REGION Network 6
   RUNG wire#powerrail
      "FB_CONCAT_STRINGS_FOR_MQTT_DB"(temperature1 := "DB_GlobalData".RTDs.RTD1.ch0, temperature2 := "DB_GlobalData".RTDs.RTD1.ch1, temperature3 := "DB_GlobalData".RTDs.RTD1.ch2, temperature4 := "DB_GlobalData".RTDs.RTD1.ch3, strCombinedString => "MQTT_DB".MQTT_CLIEENTS[0].mqttUserControl.sStringToPublish, q_aStringToSendToMqtt =>)
      "FB_CONCAT_STRINGS_FOR_MQTT_1_DB"(temperature1 := "DB_GlobalData".RTDs.RTD1.ch0, temperature2 := "DB_GlobalData".RTDs.RTD1.ch1, temperature3 :=, temperature4 := "DB_GlobalData".RTDs.RTD1.ch2, customText := '', strCombinedString =>, q_aStringToSendToMqtt => "MQTT_DB".MQTT_CLIENTS_WSTRING[0].mqttParam.message)
   END_RUNG
   // the same network as SCL:
   "FB_CONCAT_STRINGS_FOR_MQTT_DB"(temperature1 := "DB_GlobalData".RTDs.RTD1.ch0,   // "FB_CONCAT_STRINGS_FOR_MQTT"
                           temperature2 := "DB_GlobalData".RTDs.RTD1.ch1,
                           temperature3 := "DB_GlobalData".RTDs.RTD1.ch2,
                           temperature4 := "DB_GlobalData".RTDs.RTD1.ch3,
                           strCombinedString => "MQTT_DB".MQTT_CLIEENTS[0].mqttUserControl.sStringToPublish,
                           ENO => #_w1);
   IF #_w1 THEN
       "FB_CONCAT_STRINGS_FOR_MQTT_1_DB"(temperature1 := "DB_GlobalData".RTDs.RTD1.ch0,   // "FB_CONCAT_STRINGS_FOR_MQTT_1"
                               temperature2 := "DB_GlobalData".RTDs.RTD1.ch1,
                               temperature4 := "DB_GlobalData".RTDs.RTD1.ch2,
                               customText := '',
                               q_aStringToSendToMqtt => "MQTT_DB".MQTT_CLIENTS_WSTRING[0].mqttParam.message);
   END_IF;
END_REGION

REGION Network 7: MQTT publisher 1
   RUNG wire#powerrail
      "LMqtt_Publisher_DB1"(publish := wire#w1, enable := "MQTT_DB".MQTT_CLIEENTS[0].mqttUserControl.xEnable, tcpConnParam := "MQTT_DB".MQTT_CLIEENTS[0].mqttTcpParam, mqttParam := "MQTT_DB".MQTT_CLIEENTS[0].mqttParam, tcpEstablished => "MQTT_DB".MQTT_CLIEENTS[0].mqttUserControl.Status.xtcpEsablished, mqttEstablished => "MQTT_DB".MQTT_CLIEENTS[0].mqttUserControl.Status.xmqttEstavlished, published => "MQTT_DB".MQTT_CLIEENTS[0].mqttUserControl.Status.xpublished, busy => "MQTT_DB".MQTT_CLIEENTS[0].mqttUserControl.Status.xbusy, error => "MQTT_DB".MQTT_CLIEENTS[0].mqttUserControl.Status.xerror, status => "MQTT_DB".MQTT_CLIEENTS[0].mqttUserControl.Status.status, statusID => "MQTT_DB".MQTT_CLIEENTS[0].mqttUserControl.Status.istatusID)
   END_RUNG
   RUNG wire#powerrail
      Contact( "MQTT_DB".MQTT_CLIEENTS[0].mqttUserControl.xPusblish )
   END_RUNG wire#w1
   // the same network as SCL:
   "LMqtt_Publisher_DB1"(enable := "MQTT_DB".MQTT_CLIEENTS[0].mqttUserControl.xEnable,   // "LMqtt_Publisher"
                         publish := "MQTT_DB".MQTT_CLIEENTS[0].mqttUserControl.xPusblish,
                         tcpConnParam := "MQTT_DB".MQTT_CLIEENTS[0].mqttTcpParam,
                         mqttParam := "MQTT_DB".MQTT_CLIEENTS[0].mqttParam,
                         tcpEstablished => "MQTT_DB".MQTT_CLIEENTS[0].mqttUserControl.Status.xtcpEsablished,
                         mqttEstablished => "MQTT_DB".MQTT_CLIEENTS[0].mqttUserControl.Status.xmqttEstavlished,
                         published => "MQTT_DB".MQTT_CLIEENTS[0].mqttUserControl.Status.xpublished,
                         busy => "MQTT_DB".MQTT_CLIEENTS[0].mqttUserControl.Status.xbusy,
                         error => "MQTT_DB".MQTT_CLIEENTS[0].mqttUserControl.Status.xerror,
                         status => "MQTT_DB".MQTT_CLIEENTS[0].mqttUserControl.Status.status,
                         statusID => "MQTT_DB".MQTT_CLIEENTS[0].mqttUserControl.Status.istatusID);
END_REGION

REGION Network 8: MQTT-WSTRING-TEST
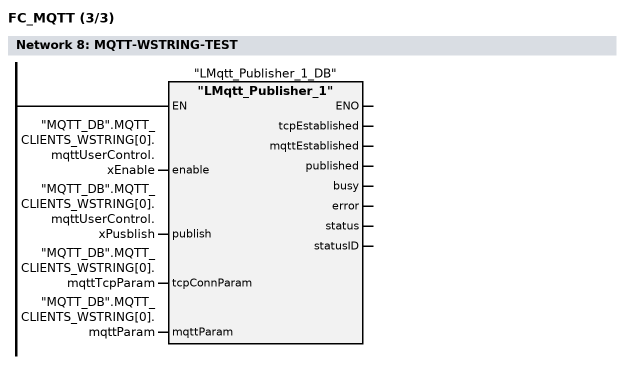
   RUNG wire#powerrail
      "LMqtt_Publisher_1_DB"(enable := "MQTT_DB".MQTT_CLIENTS_WSTRING[0].mqttUserControl.xEnable, publish := "MQTT_DB".MQTT_CLIENTS_WSTRING[0].mqttUserControl.xPusblish, tcpConnParam := "MQTT_DB".MQTT_CLIENTS_WSTRING[0].mqttTcpParam, mqttParam := "MQTT_DB".MQTT_CLIENTS_WSTRING[0].mqttParam, tcpEstablished =>, mqttEstablished =>, published =>, busy =>, error =>, status =>, statusID =>)
   END_RUNG
   // the same network as SCL:
   "LMqtt_Publisher_1_DB"(enable := "MQTT_DB".MQTT_CLIENTS_WSTRING[0].mqttUserControl.xEnable,   // "LMqtt_Publisher_1"
                          publish := "MQTT_DB".MQTT_CLIENTS_WSTRING[0].mqttUserControl.xPusblish,
                          tcpConnParam := "MQTT_DB".MQTT_CLIENTS_WSTRING[0].mqttTcpParam,
                          mqttParam := "MQTT_DB".MQTT_CLIENTS_WSTRING[0].mqttParam);
END_REGION
END_FUNCTION

FUNCTION "FC_CalculatePressRPM" : Void   // FC9, LAD
{ S7_Optimized_Access := 'TRUE' }
VERSION : 0.1
   VAR_INPUT
      i_xPulse : Bool;   // Pulse for every turn
   END_VAR
   VAR_IN_OUT
      i_iCurrentCounter : Int;
      q_iRealSPeed : Int;
   END_VAR
   VAR_TEMP
      xcalculateRPM : Bool;
      _xton : Bool;
      Temp_RPM : Real;
   END_VAR
   VAR_TEMP   // added for the SCL form of the ladder/FBD networks
      _w1 : Bool;
   END_VAR
BEGIN

REGION Network 2: 5S TIMER
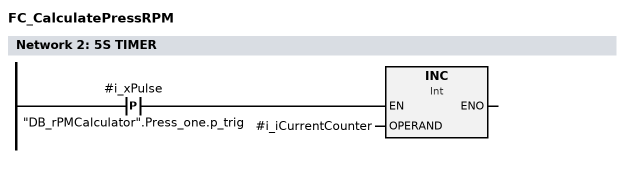
   RUNG wire#powerrail
      P_Contact(operand := #i_xPulse, bit := "DB_rPMCalculator".Press_one.p_trig)
      { S7_Templates := "DestType := Int" } Inc( #i_iCurrentCounter )
   END_RUNG
   // the same network as SCL:
   #_w1 := #i_xPulse AND NOT "DB_rPMCalculator".Press_one.p_trig;   // rising edge of #i_xPulse
   "DB_rPMCalculator".Press_one.p_trig := #i_xPulse;
   IF #_w1 THEN #i_iCurrentCounter := #i_iCurrentCounter + 1; END_IF;
END_REGION

REGION Network 3 (SCL)
   // Start 5-second timer
   "DB_rPMCalculator".Press_one.PulseTimer(IN := TRUE, PT := T#5s);



   // When 5 seconds have passed, calculate RPM
   IF "DB_rPMCalculator".Press_one.PulseTimer.Q THEN
       #q_iRealSPeed := INT_TO_REAL(#i_iCurrentCounter * 60.0) / (5.0);  // Calculate RPM
      // #q_iRealSPeed := #Temp_RPM;                      // Set the output RPM

       // Reset pulse count and timer
       #i_iCurrentCounter := 0;
       "DB_rPMCalculator".Press_one.PulseTimer(IN := FALSE,
                                               PT := T#5s);                // Reset the timer
   END_IF;
END_REGION
END_FUNCTION

FUNCTION "FC_AKD_PNU" : Void   // FC10, LAD
{ S7_Optimized_Access := 'TRUE' }
VERSION : 0.1
   VAR_INPUT
      HW_IO_telegram : Hw_Io;
   END_VAR
   VAR_IN_OUT
      AKD_PNU_v02_Instance : "AKD_PNU_v02";
      IO_DATA : "PNU_DATA";
   END_VAR
BEGIN

REGION Network 1: AKD1
   // AKD FB
   // 
   // set ID - to telegram ID of a AKD
   // 
   // 
   // # Read data from AKD PNU #
   // =================================================
   // 
   // 1. set PNU number and PNU subindex (iPNUnumber, iPNUsubindex)
   // 2. set cmd.xstartRead bit to One
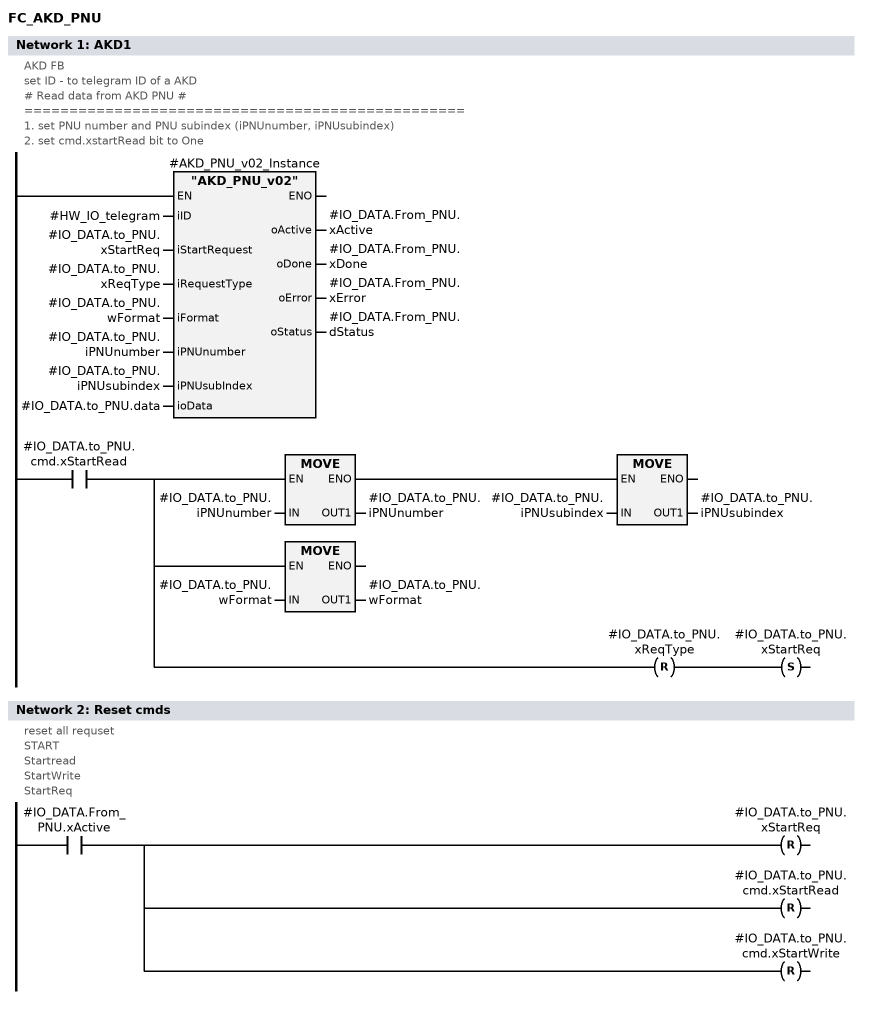
   RUNG wire#powerrail
      #AKD_PNU_v02_Instance(iID := #HW_IO_telegram, iStartRequest := #IO_DATA.to_PNU.xStartReq, iRequestType := #IO_DATA.to_PNU.xReqType, iFormat := #IO_DATA.to_PNU.wFormat, iPNUnumber := #IO_DATA.to_PNU.iPNUnumber, iPNUsubIndex := #IO_DATA.to_PNU.iPNUsubindex, ioData := #IO_DATA.to_PNU.data, oActive => #IO_DATA.From_PNU.xActive, oDone => #IO_DATA.From_PNU.xDone, oError => #IO_DATA.From_PNU.xError, oStatus => #IO_DATA.From_PNU.dStatus)
   END_RUNG
   RUNG wire#powerrail
      Contact( #IO_DATA.to_PNU.cmd.xStartRead )
      wire#w1
      Move(in := #IO_DATA.to_PNU.iPNUnumber, out1 => #IO_DATA.to_PNU.iPNUnumber)
      Move(in := #IO_DATA.to_PNU.iPNUsubindex, out1 => #IO_DATA.to_PNU.iPNUsubindex)
   END_RUNG
   RUNG wire#w1
      Move(in := #IO_DATA.to_PNU.wFormat, out1 => #IO_DATA.to_PNU.wFormat)
   END_RUNG
   RUNG wire#w1
      R_Coil( #IO_DATA.to_PNU.xReqType )
      S_Coil( #IO_DATA.to_PNU.xStartReq )
   END_RUNG
   // the same network as SCL:
   #AKD_PNU_v02_Instance(iID := #HW_IO_telegram,   // "AKD_PNU_v02"
                         iStartRequest := #IO_DATA.to_PNU.xStartReq,
                         iRequestType := #IO_DATA.to_PNU.xReqType,
                         iFormat := #IO_DATA.to_PNU.wFormat,
                         iPNUnumber := #IO_DATA.to_PNU.iPNUnumber,
                         iPNUsubIndex := #IO_DATA.to_PNU.iPNUsubindex,
                         ioData := #IO_DATA.to_PNU.data,
                         oActive => #IO_DATA.From_PNU.xActive,
                         oDone => #IO_DATA.From_PNU.xDone,
                         oError => #IO_DATA.From_PNU.xError,
                         oStatus => #IO_DATA.From_PNU.dStatus);
   IF #IO_DATA.to_PNU.cmd.xStartRead THEN
       #IO_DATA.to_PNU.iPNUnumber := #IO_DATA.to_PNU.iPNUnumber;
       #IO_DATA.to_PNU.iPNUsubindex := #IO_DATA.to_PNU.iPNUsubindex;
       #IO_DATA.to_PNU.wFormat := #IO_DATA.to_PNU.wFormat;
       #IO_DATA.to_PNU.xReqType := FALSE;
       #IO_DATA.to_PNU.xStartReq := TRUE;
   END_IF;
END_REGION

REGION Network 2: Reset cmds
   // reset all requset
   // 
   // START
   // Startread
   // StartWrite
   // StartReq
   RUNG wire#powerrail
      Contact( #IO_DATA.From_PNU.xActive )
      wire#w1
      R_Coil( #IO_DATA.to_PNU.xStartReq )
   END_RUNG
   RUNG wire#w1
      R_Coil( #IO_DATA.to_PNU.cmd.xStartRead )
   END_RUNG
   RUNG wire#w1
      R_Coil( #IO_DATA.to_PNU.cmd.xStartWrite )
   END_RUNG
   // the same network as SCL:
   IF #IO_DATA.From_PNU.xActive THEN
       #IO_DATA.to_PNU.xStartReq := FALSE;
       #IO_DATA.to_PNU.cmd.xStartRead := FALSE;
       #IO_DATA.to_PNU.cmd.xStartWrite := FALSE;
   END_IF;
END_REGION
END_FUNCTION

FUNCTION "FC_MotorControl" : Void   // FC11, LAD
{ S7_Optimized_Access := 'TRUE' }
VERSION : 0.1
   VAR_TEMP
      xM1_GoPOS2 : Bool;
      xM2_goPOS2 : Bool;
      xM3_GoPOS2 : Bool;
      xM4_GoPOS2 : Bool;
      xM5_goPOS2 : Bool;
   END_VAR
BEGIN

REGION Network 1: Cylinder CONTROL
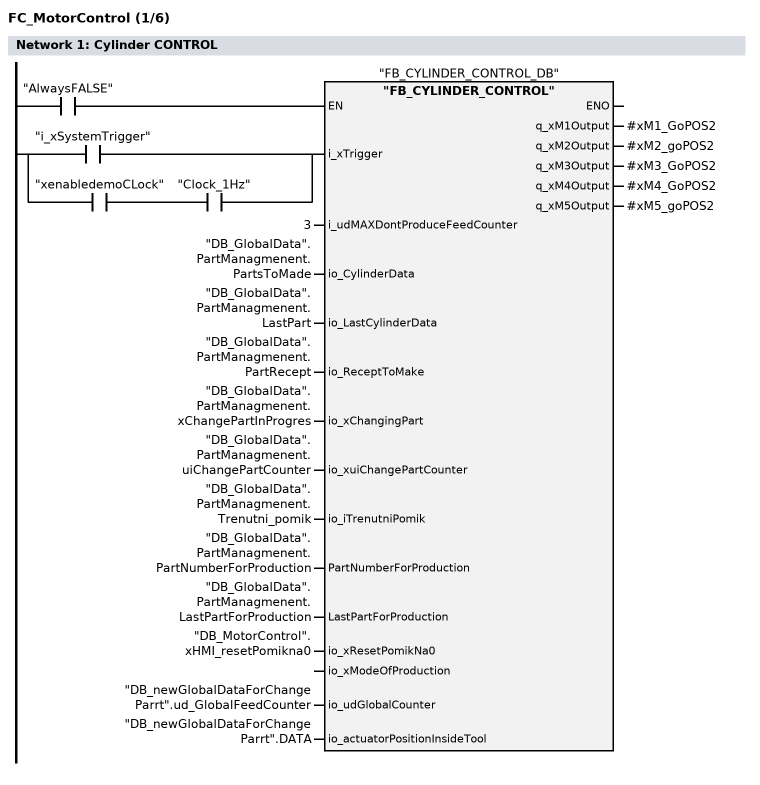
   RUNG wire#powerrail
      Contact( "AlwaysFALSE" )
      "FB_CYLINDER_CONTROL_DB"(i_xTrigger := wire#w1, i_udMAXDontProduceFeedCounter := 3, io_CylinderData := "DB_GlobalData".PartManagmenent.PartsToMade, io_LastCylinderData := "DB_GlobalData".PartManagmenent.LastPart, io_ReceptToMake := "DB_GlobalData".PartManagmenent.PartRecept, io_xChangingPart := "DB_GlobalData".PartManagmenent.xChangePartInProgres, io_xuiChangePartCounter := "DB_GlobalData".PartManagmenent.uiChangePartCounter, io_iTrenutniPomik := "DB_GlobalData".PartManagmenent.Trenutni_pomik, PartNumberForProduction := "DB_GlobalData".PartManagmenent.PartNumberForProduction, LastPartForProduction := "DB_GlobalData".PartManagmenent.LastPartForProduction, io_xResetPomikNa0 := "DB_MotorControl".xHMI_resetPomikna0, io_xModeOfProduction :=, io_udGlobalCounter := "DB_newGlobalDataForChangeParrt".ud_GlobalFeedCounter, io_actuatorPositionInsideTool := "DB_newGlobalDataForChangeParrt".DATA, q_xM1Output => #xM1_GoPOS2, q_xM2Output => #xM2_goPOS2, q_xM3Output => #xM3_GoPOS2, q_xM4Output => #xM4_GoPOS2, q_xM5Output => #xM5_goPOS2)
   END_RUNG
   RUNG wire#powerrail
      Contact( "i_xSystemTrigger" )
   END_RUNG wire#w1
   RUNG wire#powerrail
      Contact( "xenabledemoCLock" )
      Contact( "Clock_1Hz" )
   END_RUNG wire#w1
   // the same network as SCL:
   IF "AlwaysFALSE" THEN
       "FB_CYLINDER_CONTROL_DB"(i_xTrigger := "i_xSystemTrigger" OR ("xenabledemoCLock" AND "Clock_1Hz"),   // "FB_CYLINDER_CONTROL"
                               i_udMAXDontProduceFeedCounter := 3,
                               io_CylinderData := "DB_GlobalData".PartManagmenent.PartsToMade,
                               io_LastCylinderData := "DB_GlobalData".PartManagmenent.LastPart,
                               io_ReceptToMake := "DB_GlobalData".PartManagmenent.PartRecept,
                               io_xChangingPart := "DB_GlobalData".PartManagmenent.xChangePartInProgres,
                               io_xuiChangePartCounter := "DB_GlobalData".PartManagmenent.uiChangePartCounter,
                               io_iTrenutniPomik := "DB_GlobalData".PartManagmenent.Trenutni_pomik,
                               PartNumberForProduction := "DB_GlobalData".PartManagmenent.PartNumberForProduction,
                               LastPartForProduction := "DB_GlobalData".PartManagmenent.LastPartForProduction,
                               io_xResetPomikNa0 := "DB_MotorControl".xHMI_resetPomikna0,
                               io_udGlobalCounter := "DB_newGlobalDataForChangeParrt".ud_GlobalFeedCounter,
                               io_actuatorPositionInsideTool := "DB_newGlobalDataForChangeParrt".DATA,
                               q_xM1Output => #xM1_GoPOS2,
                               q_xM2Output => #xM2_goPOS2,
                               q_xM3Output => #xM3_GoPOS2,
                               q_xM4Output => #xM4_GoPOS2,
                               q_xM5Output => #xM5_goPOS2);
   END_IF;
END_REGION

REGION Network 2: Cylinde control - pipilne
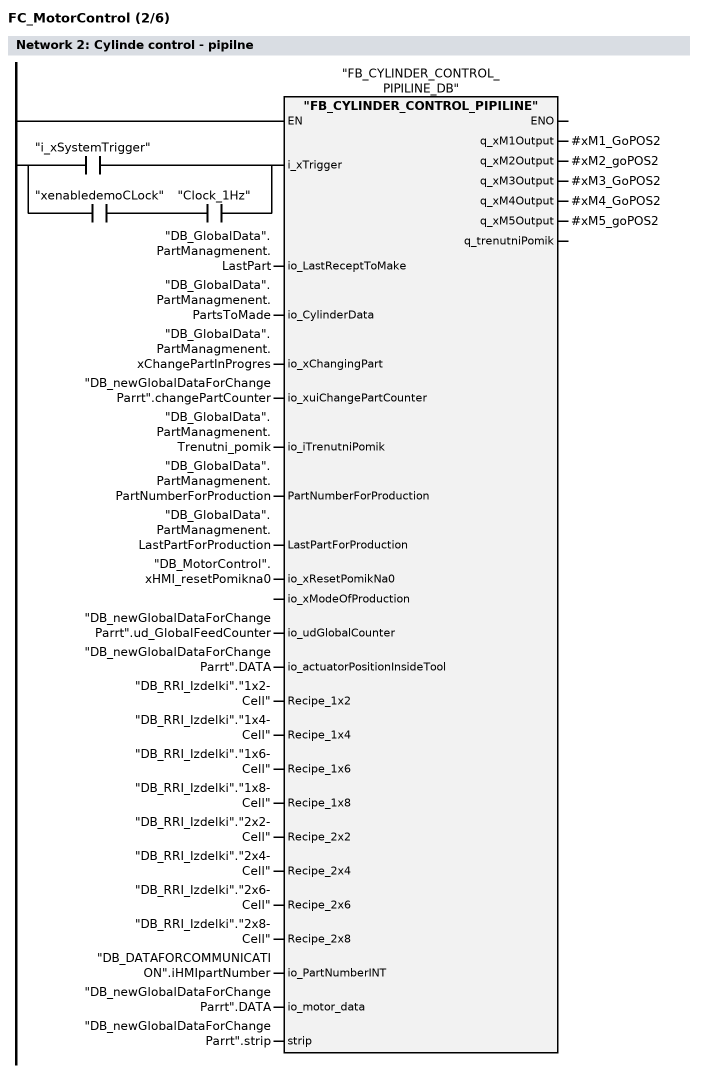
   RUNG wire#powerrail
      "FB_CYLINDER_CONTROL_PIPILINE_DB"(i_xTrigger := wire#w1, io_LastReceptToMake := "DB_GlobalData".PartManagmenent.LastPart, io_CylinderData := "DB_GlobalData".PartManagmenent.PartsToMade, io_xChangingPart := "DB_GlobalData".PartManagmenent.xChangePartInProgres, io_xuiChangePartCounter := "DB_newGlobalDataForChangeParrt".changePartCounter, io_iTrenutniPomik := "DB_GlobalData".PartManagmenent.Trenutni_pomik, PartNumberForProduction := "DB_GlobalData".PartManagmenent.PartNumberForProduction, LastPartForProduction := "DB_GlobalData".PartManagmenent.LastPartForProduction, io_xResetPomikNa0 := "DB_MotorControl".xHMI_resetPomikna0, io_xModeOfProduction :=, io_udGlobalCounter := "DB_newGlobalDataForChangeParrt".ud_GlobalFeedCounter, io_actuatorPositionInsideTool := "DB_newGlobalDataForChangeParrt".DATA, Recipe_1x2 := "DB_RRI_Izdelki"."1x2-Cell", Recipe_1x4 := "DB_RRI_Izdelki"."1x4-Cell", Recipe_1x6 := "DB_RRI_Izdelki"."1x6-Cell", Recipe_1x8 := "DB_RRI_Izdelki"."1x8-Cell", Recipe_2x2 := "DB_RRI_Izdelki"."2x2-Cell", Recipe_2x4 := "DB_RRI_Izdelki"."2x4-Cell", Recipe_2x6 := "DB_RRI_Izdelki"."2x6-Cell", Recipe_2x8 := "DB_RRI_Izdelki"."2x8-Cell", io_PartNumberINT := "DB_DATAFORCOMMUNICATION".iHMIpartNumber, io_motor_data := "DB_newGlobalDataForChangeParrt".DATA, strip := "DB_newGlobalDataForChangeParrt".strip, q_xM1Output => #xM1_GoPOS2, q_xM2Output => #xM2_goPOS2, q_xM3Output => #xM3_GoPOS2, q_xM4Output => #xM4_GoPOS2, q_xM5Output => #xM5_goPOS2, q_trenutniPomik =>)
   END_RUNG
   RUNG wire#powerrail
      Contact( "i_xSystemTrigger" )
   END_RUNG wire#w1
   RUNG wire#powerrail
      Contact( "xenabledemoCLock" )
      Contact( "Clock_1Hz" )
   END_RUNG wire#w1
   // the same network as SCL:
   "FB_CYLINDER_CONTROL_PIPILINE_DB"(i_xTrigger := "i_xSystemTrigger" OR ("xenabledemoCLock" AND "Clock_1Hz"),   // "FB_CYLINDER_CONTROL_PIPILINE"
                           io_LastReceptToMake := "DB_GlobalData".PartManagmenent.LastPart,
                           io_CylinderData := "DB_GlobalData".PartManagmenent.PartsToMade,
                           io_xChangingPart := "DB_GlobalData".PartManagmenent.xChangePartInProgres,
                           io_xuiChangePartCounter := "DB_newGlobalDataForChangeParrt".changePartCounter,
                           io_iTrenutniPomik := "DB_GlobalData".PartManagmenent.Trenutni_pomik,
                           PartNumberForProduction := "DB_GlobalData".PartManagmenent.PartNumberForProduction,
                           LastPartForProduction := "DB_GlobalData".PartManagmenent.LastPartForProduction,
                           io_xResetPomikNa0 := "DB_MotorControl".xHMI_resetPomikna0,
                           io_udGlobalCounter := "DB_newGlobalDataForChangeParrt".ud_GlobalFeedCounter,
                           io_actuatorPositionInsideTool := "DB_newGlobalDataForChangeParrt".DATA,
                           Recipe_1x2 := "DB_RRI_Izdelki"."1x2-Cell",
                           Recipe_1x4 := "DB_RRI_Izdelki"."1x4-Cell",
                           Recipe_1x6 := "DB_RRI_Izdelki"."1x6-Cell",
                           Recipe_1x8 := "DB_RRI_Izdelki"."1x8-Cell",
                           Recipe_2x2 := "DB_RRI_Izdelki"."2x2-Cell",
                           Recipe_2x4 := "DB_RRI_Izdelki"."2x4-Cell",
                           Recipe_2x6 := "DB_RRI_Izdelki"."2x6-Cell",
                           Recipe_2x8 := "DB_RRI_Izdelki"."2x8-Cell",
                           io_PartNumberINT := "DB_DATAFORCOMMUNICATION".iHMIpartNumber,
                           io_motor_data := "DB_newGlobalDataForChangeParrt".DATA,
                           strip := "DB_newGlobalDataForChangeParrt".strip,
                           q_xM1Output => #xM1_GoPOS2,
                           q_xM2Output => #xM2_goPOS2,
                           q_xM3Output => #xM3_GoPOS2,
                           q_xM4Output => #xM4_GoPOS2,
                           q_xM5Output => #xM5_goPOS2);
END_REGION

REGION Network 3
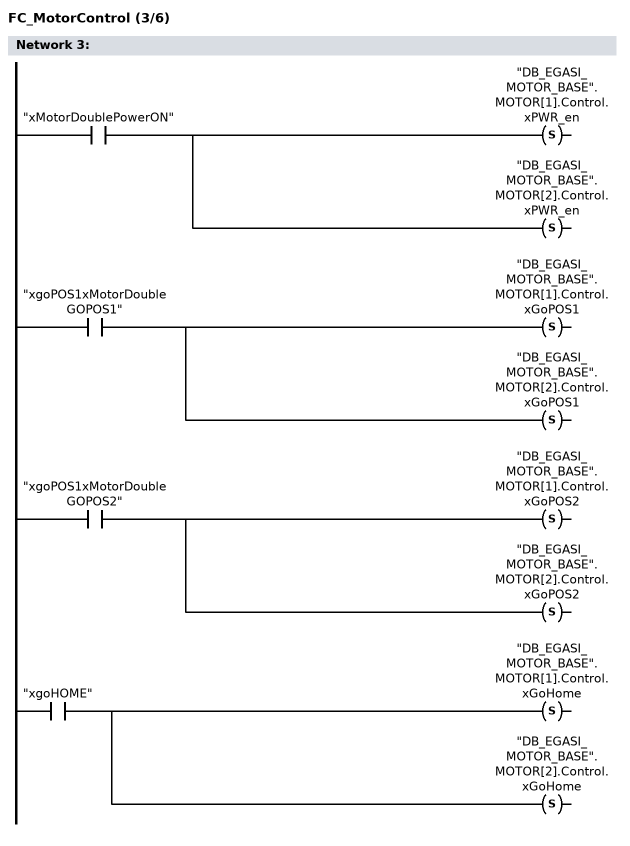
   RUNG wire#powerrail
      Contact( "xMotorDoublePowerON" )
      wire#w1
      S_Coil( "DB_EGASI_MOTOR_BASE".MOTOR[1].Control.xPWR_en )
   END_RUNG
   RUNG wire#w1
      S_Coil( "DB_EGASI_MOTOR_BASE".MOTOR[2].Control.xPWR_en )
   END_RUNG
   RUNG wire#powerrail
      Contact( "xgoPOS1xMotorDoubleGOPOS1" )
      wire#w2
      S_Coil( "DB_EGASI_MOTOR_BASE".MOTOR[1].Control.xGoPOS1 )
   END_RUNG
   RUNG wire#w2
      S_Coil( "DB_EGASI_MOTOR_BASE".MOTOR[2].Control.xGoPOS1 )
   END_RUNG
   RUNG wire#powerrail
      Contact( "xgoPOS1xMotorDoubleGOPOS2" )
      wire#w3
      S_Coil( "DB_EGASI_MOTOR_BASE".MOTOR[1].Control.xGoPOS2 )
   END_RUNG
   RUNG wire#w3
      S_Coil( "DB_EGASI_MOTOR_BASE".MOTOR[2].Control.xGoPOS2 )
   END_RUNG
   RUNG wire#powerrail
      Contact( "xgoHOME" )
      wire#w4
      S_Coil( "DB_EGASI_MOTOR_BASE".MOTOR[1].Control.xGoHome )
   END_RUNG
   RUNG wire#w4
      S_Coil( "DB_EGASI_MOTOR_BASE".MOTOR[2].Control.xGoHome )
   END_RUNG
   // the same network as SCL:
   IF "xMotorDoublePowerON" THEN
       "DB_EGASI_MOTOR_BASE".MOTOR[1].Control.xPWR_en := TRUE;
       "DB_EGASI_MOTOR_BASE".MOTOR[2].Control.xPWR_en := TRUE;
   END_IF;
   IF "xgoPOS1xMotorDoubleGOPOS1" THEN
       "DB_EGASI_MOTOR_BASE".MOTOR[1].Control.xGoPOS1 := TRUE;
       "DB_EGASI_MOTOR_BASE".MOTOR[2].Control.xGoPOS1 := TRUE;
   END_IF;
   IF "xgoPOS1xMotorDoubleGOPOS2" THEN
       "DB_EGASI_MOTOR_BASE".MOTOR[1].Control.xGoPOS2 := TRUE;
       "DB_EGASI_MOTOR_BASE".MOTOR[2].Control.xGoPOS2 := TRUE;
   END_IF;
   IF "xgoHOME" THEN
       "DB_EGASI_MOTOR_BASE".MOTOR[1].Control.xGoHome := TRUE;
       "DB_EGASI_MOTOR_BASE".MOTOR[2].Control.xGoHome := TRUE;
   END_IF;
END_REGION

REGION Network 4: EGASI MOTOR CONTROL
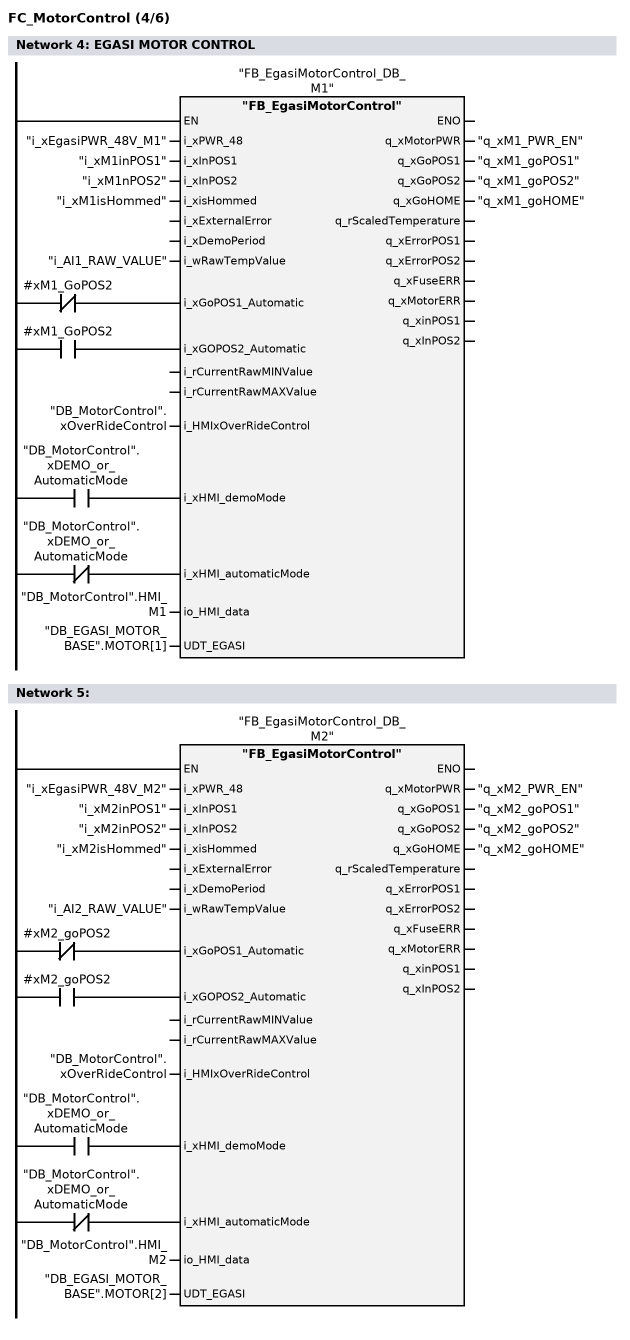
   RUNG wire#powerrail
      "FB_EgasiMotorControl_DB_M1"(i_xGoPOS1_Automatic := wire#w1, i_xGOPOS2_Automatic := wire#w2, i_xHMI_demoMode := wire#w3, i_xHMI_automaticMode := wire#w4, i_xPWR_48 := "i_xEgasiPWR_48V_M1", i_xInPOS1 := "i_xM1inPOS1", i_xInPOS2 := "i_xM1nPOS2", i_xisHommed := "i_xM1isHommed", i_xExternalError :=, i_xDemoPeriod :=, i_wRawTempValue := "i_AI1_RAW_VALUE", i_rCurrentRawMINValue :=, i_rCurrentRawMAXValue :=, i_HMIxOverRideControl := "DB_MotorControl".xOverRideControl, io_HMI_data := "DB_MotorControl".HMI_M1, UDT_EGASI := "DB_EGASI_MOTOR_BASE".MOTOR[1], q_xMotorPWR => "q_xM1_PWR_EN", q_xGoPOS1 => "q_xM1_goPOS1", q_xGoPOS2 => "q_xM1_goPOS2", q_xGoHOME => "q_xM1_goHOME", q_rScaledTemperature =>, q_xErrorPOS1 =>, q_xErrorPOS2 =>, q_xFuseERR =>, q_xMotorERR =>, q_xinPOS1 =>, q_xInPOS2 =>)
   END_RUNG
   RUNG wire#powerrail
      I_Contact( #xM1_GoPOS2 )
   END_RUNG wire#w1
   RUNG wire#powerrail
      Contact( #xM1_GoPOS2 )
   END_RUNG wire#w2
   RUNG wire#powerrail
      Contact( "DB_MotorControl".xDEMO_or_AutomaticMode )
   END_RUNG wire#w3
   RUNG wire#powerrail
      I_Contact( "DB_MotorControl".xDEMO_or_AutomaticMode )
   END_RUNG wire#w4
   // the same network as SCL:
   "FB_EgasiMotorControl_DB_M1"(i_xPWR_48 := "i_xEgasiPWR_48V_M1",   // "FB_EgasiMotorControl"
                           i_xInPOS1 := "i_xM1inPOS1",
                           i_xInPOS2 := "i_xM1nPOS2",
                           i_xisHommed := "i_xM1isHommed",
                           i_wRawTempValue := "i_AI1_RAW_VALUE",
                           i_xGoPOS1_Automatic := NOT #xM1_GoPOS2,
                           i_xGOPOS2_Automatic := #xM1_GoPOS2,
                           i_HMIxOverRideControl := "DB_MotorControl".xOverRideControl,
                           i_xHMI_demoMode := "DB_MotorControl".xDEMO_or_AutomaticMode,
                           i_xHMI_automaticMode := NOT "DB_MotorControl".xDEMO_or_AutomaticMode,
                           io_HMI_data := "DB_MotorControl".HMI_M1,
                           UDT_EGASI := "DB_EGASI_MOTOR_BASE".MOTOR[1],
                           q_xMotorPWR => "q_xM1_PWR_EN",
                           q_xGoPOS1 => "q_xM1_goPOS1",
                           q_xGoPOS2 => "q_xM1_goPOS2",
                           q_xGoHOME => "q_xM1_goHOME");
END_REGION

REGION Network 5
   RUNG wire#powerrail
      "FB_EgasiMotorControl_DB_M2"(i_xGoPOS1_Automatic := wire#w1, i_xGOPOS2_Automatic := wire#w2, i_xHMI_demoMode := wire#w3, i_xHMI_automaticMode := wire#w4, i_xPWR_48 := "i_xEgasiPWR_48V_M2", i_xInPOS1 := "i_xM2inPOS1", i_xInPOS2 := "i_xM2inPOS2", i_xisHommed := "i_xM2isHommed", i_xExternalError :=, i_xDemoPeriod :=, i_wRawTempValue := "i_AI2_RAW_VALUE", i_rCurrentRawMINValue :=, i_rCurrentRawMAXValue :=, i_HMIxOverRideControl := "DB_MotorControl".xOverRideControl, io_HMI_data := "DB_MotorControl".HMI_M2, UDT_EGASI := "DB_EGASI_MOTOR_BASE".MOTOR[2], q_xMotorPWR => "q_xM2_PWR_EN", q_xGoPOS1 => "q_xM2_goPOS1", q_xGoPOS2 => "q_xM2_goPOS2", q_xGoHOME => "q_xM2_goHOME", q_rScaledTemperature =>, q_xErrorPOS1 =>, q_xErrorPOS2 =>, q_xFuseERR =>, q_xMotorERR =>, q_xinPOS1 =>, q_xInPOS2 =>)
   END_RUNG
   RUNG wire#powerrail
      I_Contact( #xM2_goPOS2 )
   END_RUNG wire#w1
   RUNG wire#powerrail
      Contact( #xM2_goPOS2 )
   END_RUNG wire#w2
   RUNG wire#powerrail
      Contact( "DB_MotorControl".xDEMO_or_AutomaticMode )
   END_RUNG wire#w3
   RUNG wire#powerrail
      I_Contact( "DB_MotorControl".xDEMO_or_AutomaticMode )
   END_RUNG wire#w4
   // the same network as SCL:
   "FB_EgasiMotorControl_DB_M2"(i_xPWR_48 := "i_xEgasiPWR_48V_M2",   // "FB_EgasiMotorControl"
                           i_xInPOS1 := "i_xM2inPOS1",
                           i_xInPOS2 := "i_xM2inPOS2",
                           i_xisHommed := "i_xM2isHommed",
                           i_wRawTempValue := "i_AI2_RAW_VALUE",
                           i_xGoPOS1_Automatic := NOT #xM2_goPOS2,
                           i_xGOPOS2_Automatic := #xM2_goPOS2,
                           i_HMIxOverRideControl := "DB_MotorControl".xOverRideControl,
                           i_xHMI_demoMode := "DB_MotorControl".xDEMO_or_AutomaticMode,
                           i_xHMI_automaticMode := NOT "DB_MotorControl".xDEMO_or_AutomaticMode,
                           io_HMI_data := "DB_MotorControl".HMI_M2,
                           UDT_EGASI := "DB_EGASI_MOTOR_BASE".MOTOR[2],
                           q_xMotorPWR => "q_xM2_PWR_EN",
                           q_xGoPOS1 => "q_xM2_goPOS1",
                           q_xGoPOS2 => "q_xM2_goPOS2",
                           q_xGoHOME => "q_xM2_goHOME");
END_REGION

REGION Network 6
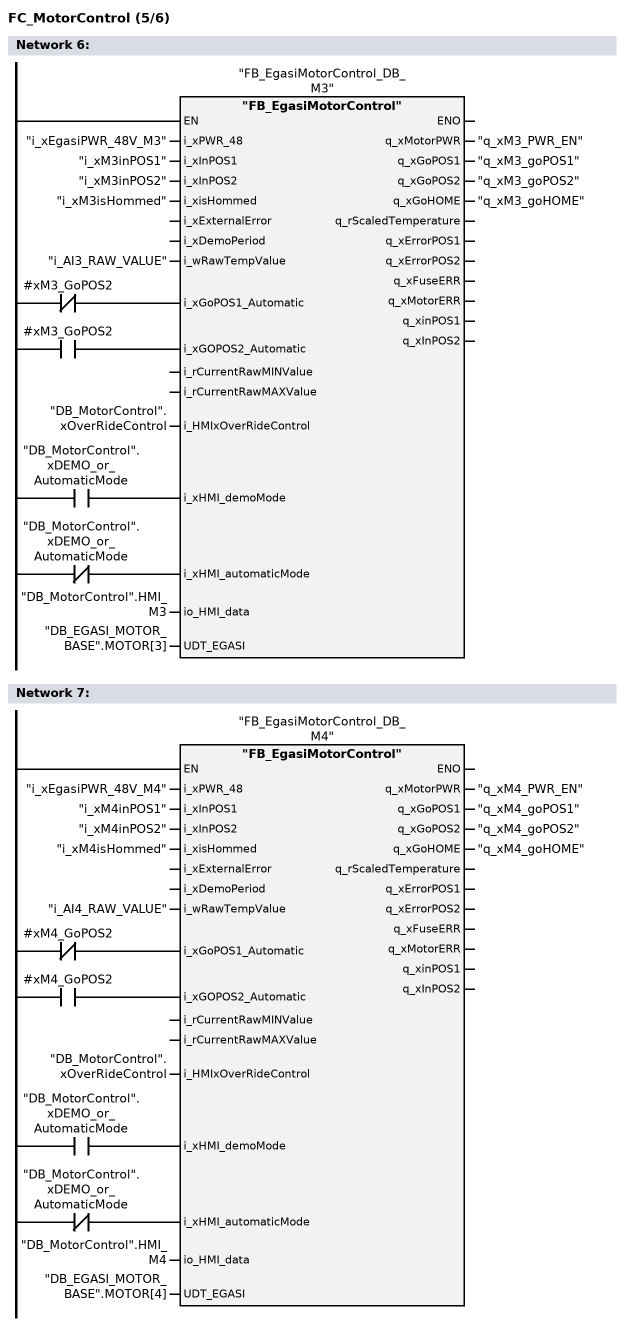
   RUNG wire#powerrail
      "FB_EgasiMotorControl_DB_M3"(i_xGoPOS1_Automatic := wire#w1, i_xGOPOS2_Automatic := wire#w2, i_xHMI_demoMode := wire#w3, i_xHMI_automaticMode := wire#w4, i_xPWR_48 := "i_xEgasiPWR_48V_M3", i_xInPOS1 := "i_xM3inPOS1", i_xInPOS2 := "i_xM3inPOS2", i_xisHommed := "i_xM3isHommed", i_xExternalError :=, i_xDemoPeriod :=, i_wRawTempValue := "i_AI3_RAW_VALUE", i_rCurrentRawMINValue :=, i_rCurrentRawMAXValue :=, i_HMIxOverRideControl := "DB_MotorControl".xOverRideControl, io_HMI_data := "DB_MotorControl".HMI_M3, UDT_EGASI := "DB_EGASI_MOTOR_BASE".MOTOR[3], q_xMotorPWR => "q_xM3_PWR_EN", q_xGoPOS1 => "q_xM3_goPOS1", q_xGoPOS2 => "q_xM3_goPOS2", q_xGoHOME => "q_xM3_goHOME", q_rScaledTemperature =>, q_xErrorPOS1 =>, q_xErrorPOS2 =>, q_xFuseERR =>, q_xMotorERR =>, q_xinPOS1 =>, q_xInPOS2 =>)
   END_RUNG
   RUNG wire#powerrail
      I_Contact( #xM3_GoPOS2 )
   END_RUNG wire#w1
   RUNG wire#powerrail
      Contact( #xM3_GoPOS2 )
   END_RUNG wire#w2
   RUNG wire#powerrail
      Contact( "DB_MotorControl".xDEMO_or_AutomaticMode )
   END_RUNG wire#w3
   RUNG wire#powerrail
      I_Contact( "DB_MotorControl".xDEMO_or_AutomaticMode )
   END_RUNG wire#w4
   // the same network as SCL:
   "FB_EgasiMotorControl_DB_M3"(i_xPWR_48 := "i_xEgasiPWR_48V_M3",   // "FB_EgasiMotorControl"
                           i_xInPOS1 := "i_xM3inPOS1",
                           i_xInPOS2 := "i_xM3inPOS2",
                           i_xisHommed := "i_xM3isHommed",
                           i_wRawTempValue := "i_AI3_RAW_VALUE",
                           i_xGoPOS1_Automatic := NOT #xM3_GoPOS2,
                           i_xGOPOS2_Automatic := #xM3_GoPOS2,
                           i_HMIxOverRideControl := "DB_MotorControl".xOverRideControl,
                           i_xHMI_demoMode := "DB_MotorControl".xDEMO_or_AutomaticMode,
                           i_xHMI_automaticMode := NOT "DB_MotorControl".xDEMO_or_AutomaticMode,
                           io_HMI_data := "DB_MotorControl".HMI_M3,
                           UDT_EGASI := "DB_EGASI_MOTOR_BASE".MOTOR[3],
                           q_xMotorPWR => "q_xM3_PWR_EN",
                           q_xGoPOS1 => "q_xM3_goPOS1",
                           q_xGoPOS2 => "q_xM3_goPOS2",
                           q_xGoHOME => "q_xM3_goHOME");
END_REGION

REGION Network 7
   RUNG wire#powerrail
      "FB_EgasiMotorControl_DB_M4"(i_xGoPOS1_Automatic := wire#w1, i_xGOPOS2_Automatic := wire#w2, i_xHMI_demoMode := wire#w3, i_xHMI_automaticMode := wire#w4, i_xPWR_48 := "i_xEgasiPWR_48V_M4", i_xInPOS1 := "i_xM4inPOS1", i_xInPOS2 := "i_xM4inPOS2", i_xisHommed := "i_xM4isHommed", i_xExternalError :=, i_xDemoPeriod :=, i_wRawTempValue := "i_AI4_RAW_VALUE", i_rCurrentRawMINValue :=, i_rCurrentRawMAXValue :=, i_HMIxOverRideControl := "DB_MotorControl".xOverRideControl, io_HMI_data := "DB_MotorControl".HMI_M4, UDT_EGASI := "DB_EGASI_MOTOR_BASE".MOTOR[4], q_xMotorPWR => "q_xM4_PWR_EN", q_xGoPOS1 => "q_xM4_goPOS1", q_xGoPOS2 => "q_xM4_goPOS2", q_xGoHOME => "q_xM4_goHOME", q_rScaledTemperature =>, q_xErrorPOS1 =>, q_xErrorPOS2 =>, q_xFuseERR =>, q_xMotorERR =>, q_xinPOS1 =>, q_xInPOS2 =>)
   END_RUNG
   RUNG wire#powerrail
      I_Contact( #xM4_GoPOS2 )
   END_RUNG wire#w1
   RUNG wire#powerrail
      Contact( #xM4_GoPOS2 )
   END_RUNG wire#w2
   RUNG wire#powerrail
      Contact( "DB_MotorControl".xDEMO_or_AutomaticMode )
   END_RUNG wire#w3
   RUNG wire#powerrail
      I_Contact( "DB_MotorControl".xDEMO_or_AutomaticMode )
   END_RUNG wire#w4
   // the same network as SCL:
   "FB_EgasiMotorControl_DB_M4"(i_xPWR_48 := "i_xEgasiPWR_48V_M4",   // "FB_EgasiMotorControl"
                           i_xInPOS1 := "i_xM4inPOS1",
                           i_xInPOS2 := "i_xM4inPOS2",
                           i_xisHommed := "i_xM4isHommed",
                           i_wRawTempValue := "i_AI4_RAW_VALUE",
                           i_xGoPOS1_Automatic := NOT #xM4_GoPOS2,
                           i_xGOPOS2_Automatic := #xM4_GoPOS2,
                           i_HMIxOverRideControl := "DB_MotorControl".xOverRideControl,
                           i_xHMI_demoMode := "DB_MotorControl".xDEMO_or_AutomaticMode,
                           i_xHMI_automaticMode := NOT "DB_MotorControl".xDEMO_or_AutomaticMode,
                           io_HMI_data := "DB_MotorControl".HMI_M4,
                           UDT_EGASI := "DB_EGASI_MOTOR_BASE".MOTOR[4],
                           q_xMotorPWR => "q_xM4_PWR_EN",
                           q_xGoPOS1 => "q_xM4_goPOS1",
                           q_xGoPOS2 => "q_xM4_goPOS2",
                           q_xGoHOME => "q_xM4_goHOME");
END_REGION

REGION Network 8